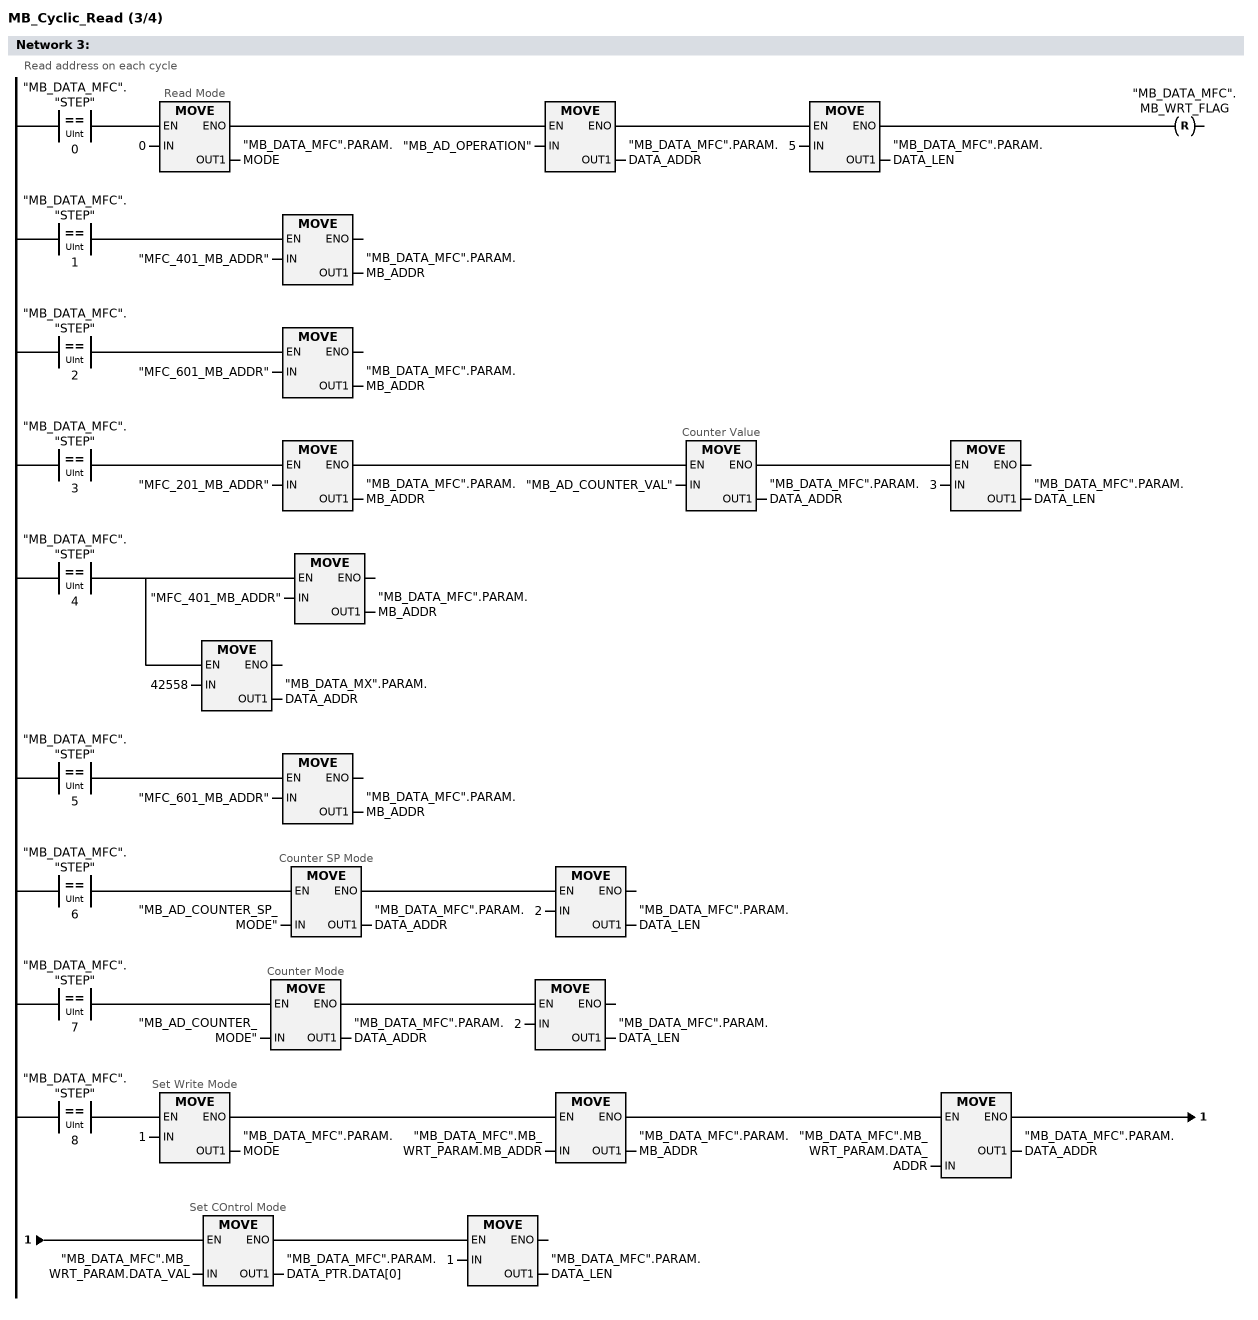
   RUNG wire#powerrail
      { S7_Templates := "SrcType := UInt" } EQ_Contact(in1 := "MB_DATA_MFC"."STEP", in2 := 0)
      Move(in := 0, out1 => "MB_DATA_MFC".PARAM.MODE)   // Read Mode
      Move(in := "MB_AD_OPERATION", out1 => "MB_DATA_MFC".PARAM.DATA_ADDR)
      Move(in := 5, out1 => "MB_DATA_MFC".PARAM.DATA_LEN)
      R_Coil( "MB_DATA_MFC".MB_WRT_FLAG )
   END_RUNG
   RUNG wire#powerrail
      { S7_Templates := "SrcType := UInt" } EQ_Contact(in1 := "MB_DATA_MFC"."STEP", in2 := 1)
      Move(in := "MFC_401_MB_ADDR", out1 => "MB_DATA_MFC".PARAM.MB_ADDR)
   END_RUNG
   RUNG wire#powerrail
      { S7_Templates := "SrcType := UInt" } EQ_Contact(in1 := "MB_DATA_MFC"."STEP", in2 := 2)
      Move(in := "MFC_601_MB_ADDR", out1 => "MB_DATA_MFC".PARAM.MB_ADDR)
   END_RUNG
   RUNG wire#powerrail
      { S7_Templates := "SrcType := UInt" } EQ_Contact(in1 := "MB_DATA_MFC"."STEP", in2 := 3)
      Move(in := "MFC_201_MB_ADDR", out1 => "MB_DATA_MFC".PARAM.MB_ADDR)
      Move(in := "MB_AD_COUNTER_VAL", out1 => "MB_DATA_MFC".PARAM.DATA_ADDR)   // Counter Value
      Move(in := 3, out1 => "MB_DATA_MFC".PARAM.DATA_LEN)
   END_RUNG
   RUNG wire#powerrail
      { S7_Templates := "SrcType := UInt" } EQ_Contact(in1 := "MB_DATA_MFC"."STEP", in2 := 4)
      wire#w1
      Move(in := "MFC_401_MB_ADDR", out1 => "MB_DATA_MFC".PARAM.MB_ADDR)
   END_RUNG
   RUNG wire#w1
      Move(in := 42558, out1 => "MB_DATA_MX".PARAM.DATA_ADDR)
   END_RUNG
   RUNG wire#powerrail
      { S7_Templates := "SrcType := UInt" } EQ_Contact(in1 := "MB_DATA_MFC"."STEP", in2 := 5)
      Move(in := "MFC_601_MB_ADDR", out1 => "MB_DATA_MFC".PARAM.MB_ADDR)
   END_RUNG
   RUNG wire#powerrail
      { S7_Templates := "SrcType := UInt" } EQ_Contact(in1 := "MB_DATA_MFC"."STEP", in2 := 6)
      Move(in := "MB_AD_COUNTER_SP_MODE", out1 => "MB_DATA_MFC".PARAM.DATA_ADDR)   // Counter SP Mode
      Move(in := 2, out1 => "MB_DATA_MFC".PARAM.DATA_LEN)
   END_RUNG
   RUNG wire#powerrail
      { S7_Templates := "SrcType := UInt" } EQ_Contact(in1 := "MB_DATA_MFC"."STEP", in2 := 7)
      Move(in := "MB_AD_COUNTER_MODE", out1 => "MB_DATA_MFC".PARAM.DATA_ADDR)   // Counter Mode
      Move(in := 2, out1 => "MB_DATA_MFC".PARAM.DATA_LEN)
   END_RUNG
   RUNG wire#powerrail
      { S7_Templates := "SrcType := UInt" } EQ_Contact(in1 := "MB_DATA_MFC"."STEP", in2 := 8)
      Move(in := 1, out1 => "MB_DATA_MFC".PARAM.MODE)   // Set Write Mode
      Move(in := "MB_DATA_MFC".MB_WRT_PARAM.MB_ADDR, out1 => "MB_DATA_MFC".PARAM.MB_ADDR)
      Move(in := "MB_DATA_MFC".MB_WRT_PARAM.DATA_ADDR, out1 => "MB_DATA_MFC".PARAM.DATA_ADDR)
      Move(in := "MB_DATA_MFC".MB_WRT_PARAM.DATA_VAL, out1 => "MB_DATA_MFC".PARAM.DATA_PTR.DATA[0])   // Set COntrol Mode
      Move(in := 1, out1 => "MB_DATA_MFC".PARAM.DATA_LEN)
   END_RUNG
   // the same network as SCL:
   IF "MB_DATA_MFC"."STEP" = 0 THEN
       "MB_DATA_MFC".PARAM.MODE := 0;   // Read Mode
       "MB_DATA_MFC".PARAM.DATA_ADDR := "MB_AD_OPERATION";
       "MB_DATA_MFC".PARAM.DATA_LEN := 5;
       "MB_DATA_MFC".MB_WRT_FLAG := FALSE;
   END_IF;
   IF "MB_DATA_MFC"."STEP" = 1 THEN "MB_DATA_MFC".PARAM.MB_ADDR := "MFC_401_MB_ADDR"; END_IF;
   IF "MB_DATA_MFC"."STEP" = 2 THEN "MB_DATA_MFC".PARAM.MB_ADDR := "MFC_601_MB_ADDR"; END_IF;
   IF "MB_DATA_MFC"."STEP" = 3 THEN
       "MB_DATA_MFC".PARAM.MB_ADDR := "MFC_201_MB_ADDR";
       "MB_DATA_MFC".PARAM.DATA_ADDR := "MB_AD_COUNTER_VAL";   // Counter Value
       "MB_DATA_MFC".PARAM.DATA_LEN := 3;
   END_IF;
   IF "MB_DATA_MFC"."STEP" = 4 THEN
       "MB_DATA_MFC".PARAM.MB_ADDR := "MFC_401_MB_ADDR";
       "MB_DATA_MX".PARAM.DATA_ADDR := 42558;
   END_IF;
   IF "MB_DATA_MFC"."STEP" = 5 THEN "MB_DATA_MFC".PARAM.MB_ADDR := "MFC_601_MB_ADDR"; END_IF;
   IF "MB_DATA_MFC"."STEP" = 6 THEN
       "MB_DATA_MFC".PARAM.DATA_ADDR := "MB_AD_COUNTER_SP_MODE";   // Counter SP Mode
       "MB_DATA_MFC".PARAM.DATA_LEN := 2;
   END_IF;
   IF "MB_DATA_MFC"."STEP" = 7 THEN
       "MB_DATA_MFC".PARAM.DATA_ADDR := "MB_AD_COUNTER_MODE";   // Counter Mode
       "MB_DATA_MFC".PARAM.DATA_LEN := 2;
   END_IF;
   IF "MB_DATA_MFC"."STEP" = 8 THEN
       "MB_DATA_MFC".PARAM.MODE := 1;   // Set Write Mode
       "MB_DATA_MFC".PARAM.MB_ADDR := "MB_DATA_MFC".MB_WRT_PARAM.MB_ADDR;
       "MB_DATA_MFC".PARAM.DATA_ADDR := "MB_DATA_MFC".MB_WRT_PARAM.DATA_ADDR;
       "MB_DATA_MFC".PARAM.DATA_PTR.DATA[0] := "MB_DATA_MFC".MB_WRT_PARAM.DATA_VAL;   // Set COntrol Mode
       "MB_DATA_MFC".PARAM.DATA_LEN := 1;
   END_IF;
END_REGION

REGION Network 4
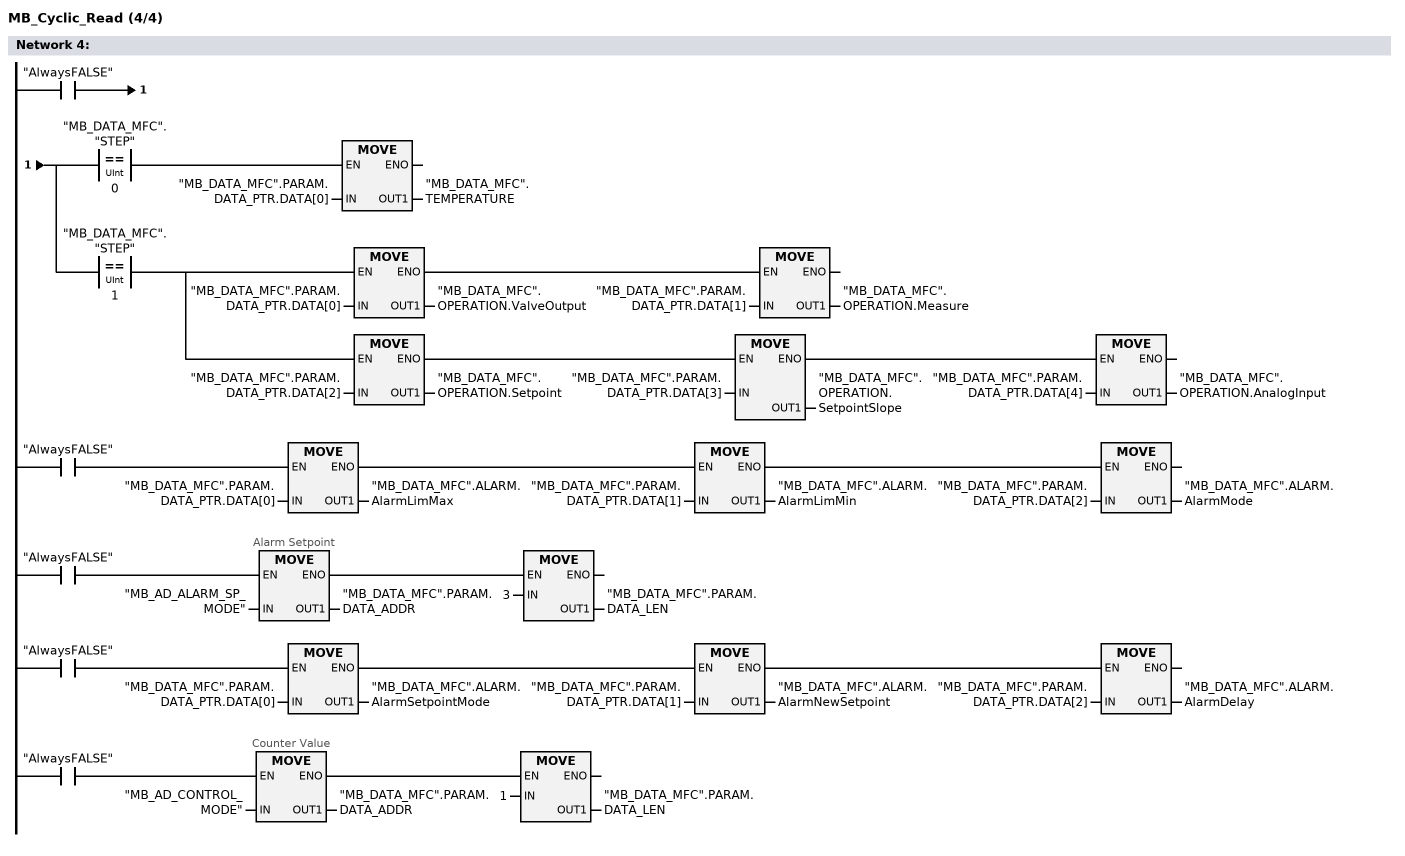
   RUNG wire#powerrail
      Contact( "AlwaysFALSE" )
      wire#w1
      { S7_Templates := "SrcType := UInt" } EQ_Contact(in1 := "MB_DATA_MFC"."STEP", in2 := 0)
      Move(in := "MB_DATA_MFC".PARAM.DATA_PTR.DATA[0], out1 => "MB_DATA_MFC".TEMPERATURE)
   END_RUNG
   RUNG wire#w1
      { S7_Templates := "SrcType := UInt" } EQ_Contact(in1 := "MB_DATA_MFC"."STEP", in2 := 1)
      wire#w2
      Move(in := "MB_DATA_MFC".PARAM.DATA_PTR.DATA[0], out1 => "MB_DATA_MFC".OPERATION.ValveOutput)
      Move(in := "MB_DATA_MFC".PARAM.DATA_PTR.DATA[1], out1 => "MB_DATA_MFC".OPERATION.Measure)
   END_RUNG
   RUNG wire#w2
      Move(in := "MB_DATA_MFC".PARAM.DATA_PTR.DATA[2], out1 => "MB_DATA_MFC".OPERATION.Setpoint)
      Move(in := "MB_DATA_MFC".PARAM.DATA_PTR.DATA[3], out1 => "MB_DATA_MFC".OPERATION.SetpointSlope)
      Move(in := "MB_DATA_MFC".PARAM.DATA_PTR.DATA[4], out1 => "MB_DATA_MFC".OPERATION.AnalogInput)
   END_RUNG
   RUNG wire#powerrail
      Contact( "AlwaysFALSE" )
      Move(in := "MB_DATA_MFC".PARAM.DATA_PTR.DATA[0], out1 => "MB_DATA_MFC".ALARM.AlarmLimMax)
      Move(in := "MB_DATA_MFC".PARAM.DATA_PTR.DATA[1], out1 => "MB_DATA_MFC".ALARM.AlarmLimMin)
      Move(in := "MB_DATA_MFC".PARAM.DATA_PTR.DATA[2], out1 => "MB_DATA_MFC".ALARM.AlarmMode)
   END_RUNG
   RUNG wire#powerrail
      Contact( "AlwaysFALSE" )
      Move(in := "MB_AD_ALARM_SP_MODE", out1 => "MB_DATA_MFC".PARAM.DATA_ADDR)   // Alarm Setpoint
      Move(in := 3, out1 => "MB_DATA_MFC".PARAM.DATA_LEN)
   END_RUNG
   RUNG wire#powerrail
      Contact( "AlwaysFALSE" )
      Move(in := "MB_DATA_MFC".PARAM.DATA_PTR.DATA[0], out1 => "MB_DATA_MFC".ALARM.AlarmSetpointMode)
      Move(in := "MB_DATA_MFC".PARAM.DATA_PTR.DATA[1], out1 => "MB_DATA_MFC".ALARM.AlarmNewSetpoint)
      Move(in := "MB_DATA_MFC".PARAM.DATA_PTR.DATA[2], out1 => "MB_DATA_MFC".ALARM.AlarmDelay)
   END_RUNG
   RUNG wire#powerrail
      Contact( "AlwaysFALSE" )
      Move(in := "MB_AD_CONTROL_MODE", out1 => "MB_DATA_MFC".PARAM.DATA_ADDR)   // Counter Value
      Move(in := 1, out1 => "MB_DATA_MFC".PARAM.DATA_LEN)
   END_RUNG
   // the same network as SCL:
   IF "AlwaysFALSE" AND ("MB_DATA_MFC"."STEP" = 0) THEN
       "MB_DATA_MFC".TEMPERATURE := "MB_DATA_MFC".PARAM.DATA_PTR.DATA[0];
   END_IF;
   IF "AlwaysFALSE" AND ("MB_DATA_MFC"."STEP" = 1) THEN
       "MB_DATA_MFC".OPERATION.ValveOutput := "MB_DATA_MFC".PARAM.DATA_PTR.DATA[0];
       "MB_DATA_MFC".OPERATION.Measure := "MB_DATA_MFC".PARAM.DATA_PTR.DATA[1];
       "MB_DATA_MFC".OPERATION.Setpoint := "MB_DATA_MFC".PARAM.DATA_PTR.DATA[2];
       "MB_DATA_MFC".OPERATION.SetpointSlope := "MB_DATA_MFC".PARAM.DATA_PTR.DATA[3];
       "MB_DATA_MFC".OPERATION.AnalogInput := "MB_DATA_MFC".PARAM.DATA_PTR.DATA[4];
   END_IF;
   IF "AlwaysFALSE" THEN
       "MB_DATA_MFC".ALARM.AlarmLimMax := "MB_DATA_MFC".PARAM.DATA_PTR.DATA[0];
       "MB_DATA_MFC".ALARM.AlarmLimMin := "MB_DATA_MFC".PARAM.DATA_PTR.DATA[1];
       "MB_DATA_MFC".ALARM.AlarmMode := "MB_DATA_MFC".PARAM.DATA_PTR.DATA[2];
       "MB_DATA_MFC".PARAM.DATA_ADDR := "MB_AD_ALARM_SP_MODE";   // Alarm Setpoint
       "MB_DATA_MFC".PARAM.DATA_LEN := 3;
       "MB_DATA_MFC".ALARM.AlarmSetpointMode := "MB_DATA_MFC".PARAM.DATA_PTR.DATA[0];
       "MB_DATA_MFC".ALARM.AlarmNewSetpoint := "MB_DATA_MFC".PARAM.DATA_PTR.DATA[1];
       "MB_DATA_MFC".ALARM.AlarmDelay := "MB_DATA_MFC".PARAM.DATA_PTR.DATA[2];
       "MB_DATA_MFC".PARAM.DATA_ADDR := "MB_AD_CONTROL_MODE";   // Counter Value
       "MB_DATA_MFC".PARAM.DATA_LEN := 1;
   END_IF;
END_REGION
END_FUNCTION

FUNCTION "TESTS_1" : Void   // FC13, LAD
{ S7_Optimized_Access := 'FALSE' }
VERSION : 0.1
   VAR_TEMP   // added for the SCL form of the ladder/FBD networks
      _w1 : Bool;
   END_VAR
BEGIN

REGION Network 1
   // ALARM Settings
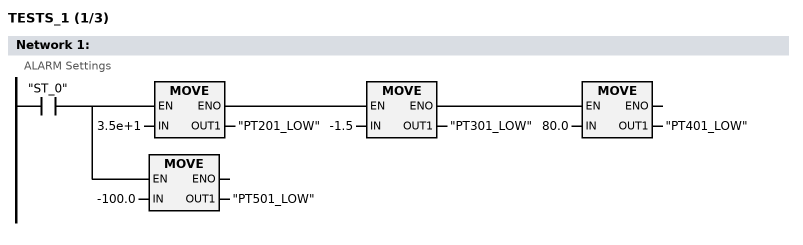
   RUNG wire#powerrail
      Contact( "ST_0" )
      wire#w1
      { S7_GenerateENO := "TRUE" } Move(in := 3.5e+1, out1 => "PT201_LOW")
      { S7_GenerateENO := "TRUE" } Move(in := -1.5, out1 => "PT301_LOW")
      { S7_GenerateENO := "TRUE" } Move(in := 80.0, out1 => "PT401_LOW")
   END_RUNG
   RUNG wire#w1
      { S7_GenerateENO := "TRUE" } Move(in := -100.0, out1 => "PT501_LOW")
   END_RUNG
   // the same network as SCL:
   // ENO of a box is taken as its EN; it also drops when the box reports an error
   IF "ST_0" THEN
       "PT201_LOW" := 3.5e+1;
       "PT301_LOW" := -1.5;
       "PT401_LOW" := 80.0;
       "PT501_LOW" := -100.0;
   END_IF;
END_REGION

REGION Network 2: Pneumatic Tests
   // Test Pneumatic System (Test #1-#6)
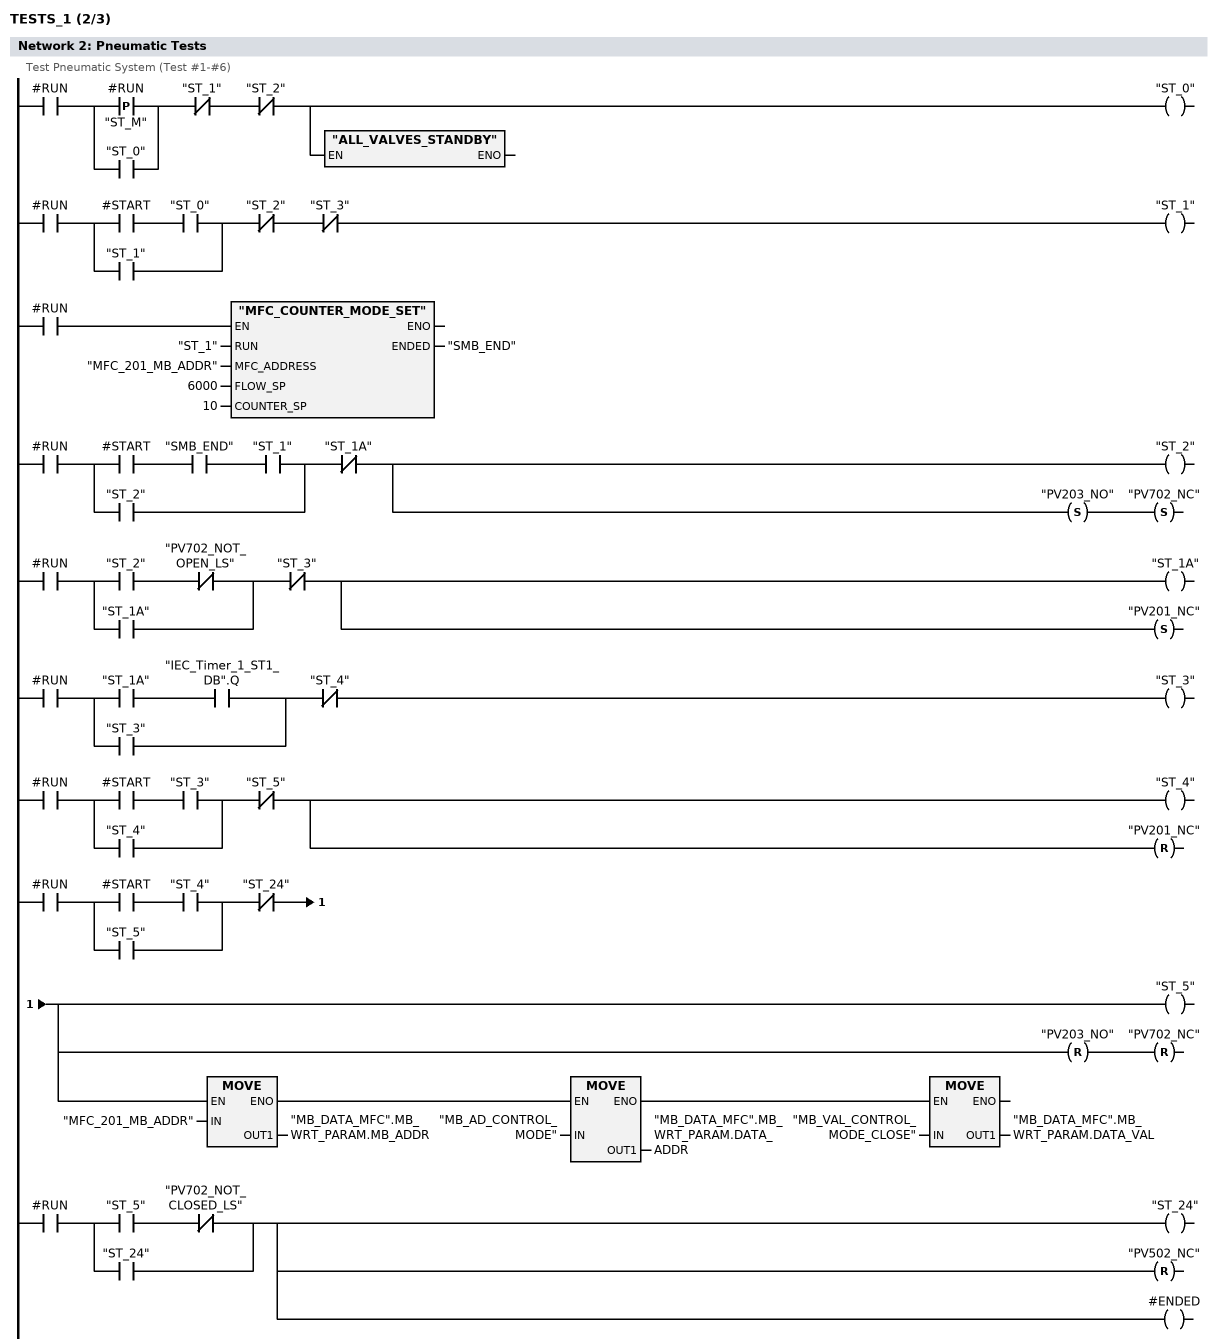
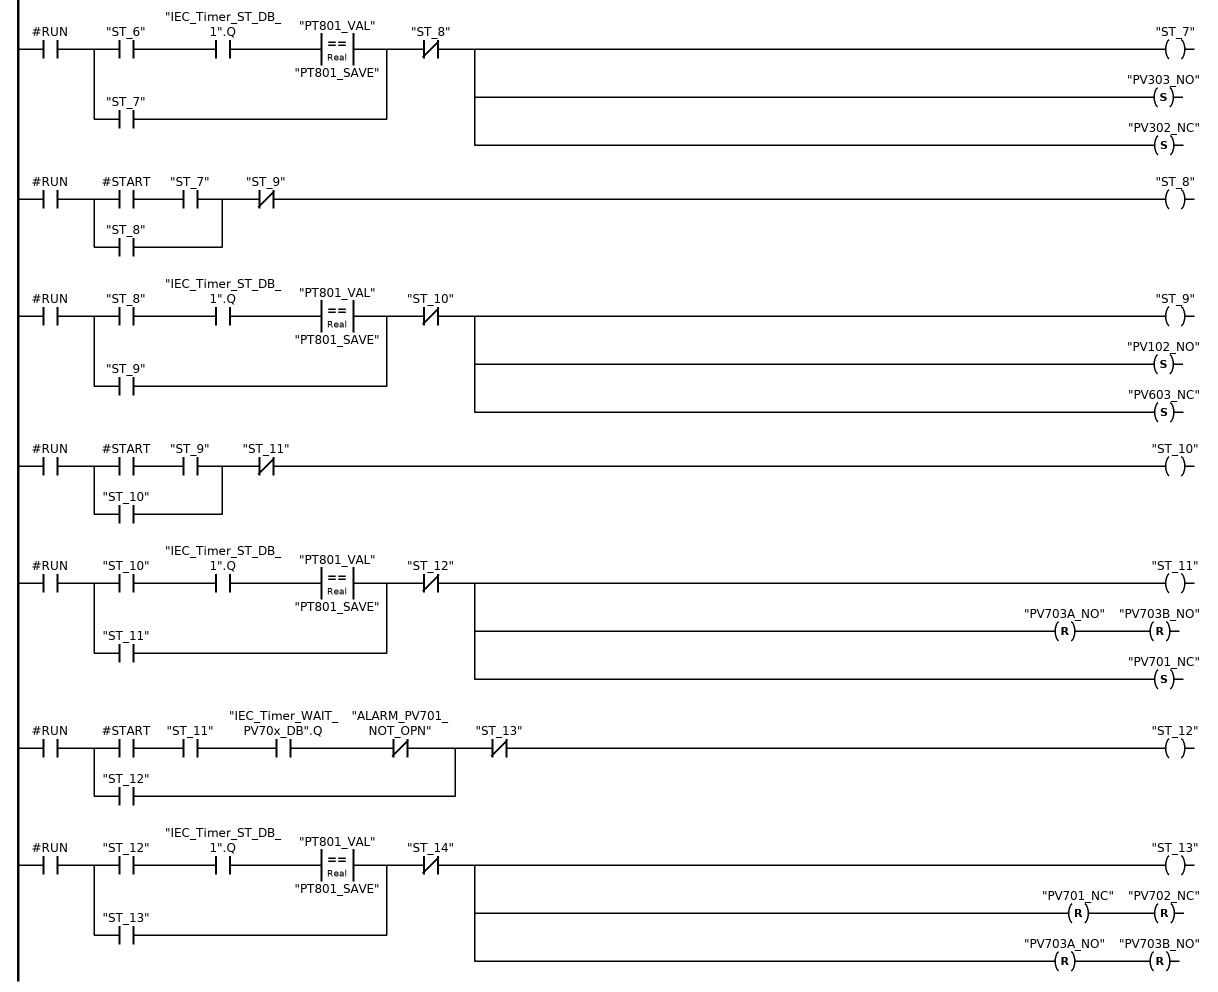
   RUNG wire#powerrail
      Contact( #RUN )
      wire#w1
      P_Contact(operand := #RUN, bit := "ST_M")
      wire#w2
      I_Contact( "ST_1" )
      I_Contact( "ST_2" )
      wire#w3
      Coil( "ST_0" )
   END_RUNG
   RUNG wire#w1
      Contact( "ST_0" )
   END_RUNG wire#w2
   RUNG wire#w3
      "ALL_VALVES_STANDBY"()
   END_RUNG
   RUNG wire#powerrail
      Contact( #RUN )
      wire#w4
      Contact( #START )
      Contact( "ST_0" )
      wire#w5
      I_Contact( "ST_2" )
      I_Contact( "ST_3" )
      Coil( "ST_1" )
   END_RUNG
   RUNG wire#w4
      Contact( "ST_1" )
   END_RUNG wire#w5
   RUNG wire#powerrail
      Contact( #RUN )
      "MFC_COUNTER_MODE_SET"(RUN := "ST_1", MFC_ADDRESS := "MFC_201_MB_ADDR", FLOW_SP := 6000, COUNTER_SP := 10, ENDED => "SMB_END")
   END_RUNG
   RUNG wire#powerrail
      Contact( #RUN )
      wire#w6
      Contact( #START )
      Contact( "SMB_END" )
      Contact( "ST_1" )
      wire#w7
      I_Contact( "ST_1A" )
      wire#w8
      Coil( "ST_2" )
   END_RUNG
   RUNG wire#w6
      Contact( "ST_2" )
   END_RUNG wire#w7
   RUNG wire#w8
      S_Coil( "PV203_NO" )
      S_Coil( "PV702_NC" )
   END_RUNG
   RUNG wire#powerrail
      Contact( #RUN )
      wire#w9
      Contact( "ST_2" )
      I_Contact( "PV702_NOT_OPEN_LS" )
      wire#w10
      I_Contact( "ST_3" )
      wire#w11
      Coil( "ST_1A" )
   END_RUNG
   RUNG wire#w9
      Contact( "ST_1A" )
   END_RUNG wire#w10
   RUNG wire#w11
      S_Coil( "PV201_NC" )
   END_RUNG
   RUNG wire#powerrail
      Contact( #RUN )
      wire#w12
      Contact( "ST_1A" )
      Contact( "IEC_Timer_1_ST1_DB".Q )
      wire#w13
      I_Contact( "ST_4" )
      Coil( "ST_3" )
   END_RUNG
   RUNG wire#w12
      Contact( "ST_3" )
   END_RUNG wire#w13
   RUNG wire#powerrail
      Contact( #RUN )
      wire#w14
      Contact( #START )
      Contact( "ST_3" )
      wire#w15
      I_Contact( "ST_5" )
      wire#w16
      Coil( "ST_4" )
   END_RUNG
   RUNG wire#w14
      Contact( "ST_4" )
   END_RUNG wire#w15
   RUNG wire#w16
      R_Coil( "PV201_NC" )
   END_RUNG
   RUNG wire#powerrail
      Contact( #RUN )
      wire#w17
      Contact( #START )
      Contact( "ST_4" )
      wire#w18
      I_Contact( "ST_24" )
      wire#w19
      Coil( "ST_5" )
   END_RUNG
   RUNG wire#w17
      Contact( "ST_5" )
   END_RUNG wire#w18
   RUNG wire#w19
      R_Coil( "PV203_NO" )
      R_Coil( "PV702_NC" )
   END_RUNG
   RUNG wire#w19
      Move(in := "MFC_201_MB_ADDR", out1 => "MB_DATA_MFC".MB_WRT_PARAM.MB_ADDR)
      Move(in := "MB_AD_CONTROL_MODE", out1 => "MB_DATA_MFC".MB_WRT_PARAM.DATA_ADDR)
      Move(in := "MB_VAL_CONTROL_MODE_CLOSE", out1 => "MB_DATA_MFC".MB_WRT_PARAM.DATA_VAL)
   END_RUNG
   RUNG wire#powerrail
      Contact( #RUN )
      wire#w20
      Contact( "ST_5" )
      I_Contact( "PV702_NOT_CLOSED_LS" )
      wire#w21
      Coil( "ST_24" )
   END_RUNG
   RUNG wire#w20
      Contact( "ST_24" )
   END_RUNG wire#w21
   RUNG wire#w21
      R_Coil( "PV502_NC" )
   END_RUNG
   RUNG wire#w21
      Coil( #ENDED )
   END_RUNG
   RUNG wire#powerrail
      Contact( #RUN )
      wire#w22
      Contact( "ST_6" )
      Contact( "IEC_Timer_ST_DB_1".Q )
      { S7_Templates := "SrcType := Real" } EQ_Contact(in1 := "PT801_VAL", in2 := "PT801_SAVE")
      wire#w23
      I_Contact( "ST_8" )
      wire#w24
      Coil( "ST_7" )
   END_RUNG
   RUNG wire#w22
      Contact( "ST_7" )
   END_RUNG wire#w23
   RUNG wire#w24
      S_Coil( "PV303_NO" )
   END_RUNG
   RUNG wire#w24
      S_Coil( "PV302_NC" )
   END_RUNG
   RUNG wire#powerrail
      Contact( #RUN )
      wire#w25
      Contact( #START )
      Contact( "ST_7" )
      wire#w26
      I_Contact( "ST_9" )
      Coil( "ST_8" )
   END_RUNG
   RUNG wire#w25
      Contact( "ST_8" )
   END_RUNG wire#w26
   RUNG wire#powerrail
      Contact( #RUN )
      wire#w27
      Contact( "ST_8" )
      Contact( "IEC_Timer_ST_DB_1".Q )
      { S7_Templates := "SrcType := Real" } EQ_Contact(in1 := "PT801_VAL", in2 := "PT801_SAVE")
      wire#w28
      I_Contact( "ST_10" )
      wire#w29
      Coil( "ST_9" )
   END_RUNG
   RUNG wire#w27
      Contact( "ST_9" )
   END_RUNG wire#w28
   RUNG wire#w29
      S_Coil( "PV102_NO" )
   END_RUNG
   RUNG wire#w29
      S_Coil( "PV603_NC" )
   END_RUNG
   RUNG wire#powerrail
      Contact( #RUN )
      wire#w30
      Contact( #START )
      Contact( "ST_9" )
      wire#w31
      I_Contact( "ST_11" )
      Coil( "ST_10" )
   END_RUNG
   RUNG wire#w30
      Contact( "ST_10" )
   END_RUNG wire#w31
   RUNG wire#powerrail
      Contact( #RUN )
      wire#w32
      Contact( "ST_10" )
      Contact( "IEC_Timer_ST_DB_1".Q )
      { S7_Templates := "SrcType := Real" } EQ_Contact(in1 := "PT801_VAL", in2 := "PT801_SAVE")
      wire#w33
      I_Contact( "ST_12" )
      wire#w34
      Coil( "ST_11" )
   END_RUNG
   RUNG wire#w32
      Contact( "ST_11" )
   END_RUNG wire#w33
   RUNG wire#w34
      R_Coil( "PV703A_NO" )
      R_Coil( "PV703B_NO" )
   END_RUNG
   RUNG wire#w34
      S_Coil( "PV701_NC" )
   END_RUNG
   RUNG wire#powerrail
      Contact( #RUN )
      wire#w35
      Contact( #START )
      Contact( "ST_11" )
      Contact( "IEC_Timer_WAIT_PV70x_DB".Q )
      I_Contact( "ALARM_PV701_NOT_OPN" )
      wire#w36
      I_Contact( "ST_13" )
      Coil( "ST_12" )
   END_RUNG
   RUNG wire#w35
      Contact( "ST_12" )
   END_RUNG wire#w36
   RUNG wire#powerrail
      Contact( #RUN )
      wire#w37
      Contact( "ST_12" )
      Contact( "IEC_Timer_ST_DB_1".Q )
      { S7_Templates := "SrcType := Real" } EQ_Contact(in1 := "PT801_VAL", in2 := "PT801_SAVE")
      wire#w38
      I_Contact( "ST_14" )
      wire#w39
      Coil( "ST_13" )
   END_RUNG
   RUNG wire#w37
      Contact( "ST_13" )
   END_RUNG wire#w38
   RUNG wire#w39
      R_Coil( "PV701_NC" )
      R_Coil( "PV702_NC" )
   END_RUNG
   RUNG wire#w39
      R_Coil( "PV703A_NO" )
      R_Coil( "PV703B_NO" )
   END_RUNG
   // the same network as SCL:
   #_w1 := #RUN AND #RUN AND NOT "ST_M";   // rising edge of #RUN
   "ST_M" := #RUN;
   "ST_0" := (#_w1 OR (#RUN AND "ST_0")) AND NOT "ST_1" AND NOT "ST_2";
   IF "ST_0" THEN "ALL_VALVES_STANDBY"(); END_IF;
   "ST_1" := #RUN AND ((#START AND "ST_0") OR "ST_1") AND NOT "ST_2" AND NOT "ST_3";
   IF #RUN THEN
       "MFC_COUNTER_MODE_SET"(RUN := "ST_1",
                              MFC_ADDRESS := "MFC_201_MB_ADDR",
                              FLOW_SP := 6000,
                              COUNTER_SP := 10,
                              ENDED => "SMB_END");
   END_IF;
   "ST_2" := #RUN AND ((#START AND "SMB_END" AND "ST_1") OR "ST_2") AND NOT "ST_1A";
   IF "ST_2" THEN
       "PV203_NO" := TRUE;
       "PV702_NC" := TRUE;
   END_IF;
   "ST_1A" := #RUN AND (("ST_2" AND NOT "PV702_NOT_OPEN_LS") OR "ST_1A") AND NOT "ST_3";
   IF "ST_1A" THEN "PV201_NC" := TRUE; END_IF;
   "ST_3" := #RUN AND (("ST_1A" AND "IEC_Timer_1_ST1_DB".Q) OR "ST_3") AND NOT "ST_4";
   "ST_4" := #RUN AND ((#START AND "ST_3") OR "ST_4") AND NOT "ST_5";
   IF "ST_4" THEN "PV201_NC" := FALSE; END_IF;
   "ST_5" := #RUN AND ((#START AND "ST_4") OR "ST_5") AND NOT "ST_24";
   IF "ST_5" THEN
       "PV203_NO" := FALSE;
       "PV702_NC" := FALSE;
       "MB_DATA_MFC".MB_WRT_PARAM.MB_ADDR := "MFC_201_MB_ADDR";
       "MB_DATA_MFC".MB_WRT_PARAM.DATA_ADDR := "MB_AD_CONTROL_MODE";
       "MB_DATA_MFC".MB_WRT_PARAM.DATA_VAL := "MB_VAL_CONTROL_MODE_CLOSE";
   END_IF;
   "ST_24" := #RUN AND (("ST_5" AND NOT "PV702_NOT_CLOSED_LS") OR "ST_24");
   IF "ST_24" THEN "PV502_NC" := FALSE; END_IF;
   #ENDED := "ST_24";
   "ST_7" := #RUN AND (("ST_6" AND "IEC_Timer_ST_DB_1".Q AND ("PT801_VAL" = "PT801_SAVE")) OR "ST_7") AND NOT "ST_8";
   IF "ST_7" THEN
       "PV303_NO" := TRUE;
       "PV302_NC" := TRUE;
   END_IF;
   "ST_8" := #RUN AND ((#START AND "ST_7") OR "ST_8") AND NOT "ST_9";
   "ST_9" := #RUN AND (("ST_8" AND "IEC_Timer_ST_DB_1".Q AND ("PT801_VAL" = "PT801_SAVE")) OR "ST_9") AND NOT "ST_10";
   IF "ST_9" THEN
       "PV102_NO" := TRUE;
       "PV603_NC" := TRUE;
   END_IF;
   "ST_10" := #RUN AND ((#START AND "ST_9") OR "ST_10") AND NOT "ST_11";
   "ST_11" := #RUN AND (("ST_10" AND "IEC_Timer_ST_DB_1".Q AND ("PT801_VAL" = "PT801_SAVE")) OR "ST_11") AND NOT "ST_12";
   IF "ST_11" THEN
       "PV703A_NO" := FALSE;
       "PV703B_NO" := FALSE;
       "PV701_NC" := TRUE;
   END_IF;
   "ST_12" := #RUN AND ((#START AND "ST_11" AND "IEC_Timer_WAIT_PV70x_DB".Q AND NOT "ALARM_PV701_NOT_OPN") OR "ST_12") AND NOT "ST_13";
   "ST_13" := #RUN AND (("ST_12" AND "IEC_Timer_ST_DB_1".Q AND ("PT801_VAL" = "PT801_SAVE")) OR "ST_13") AND NOT "ST_14";
   IF "ST_13" THEN
       "PV701_NC" := FALSE;
       "PV702_NC" := FALSE;
       "PV703A_NO" := FALSE;
       "PV703B_NO" := FALSE;
   END_IF;
END_REGION

REGION Network 3: Process Tests
   // Tests Process Circuits  (Test #7-#9)
END_REGION

REGION Network 4
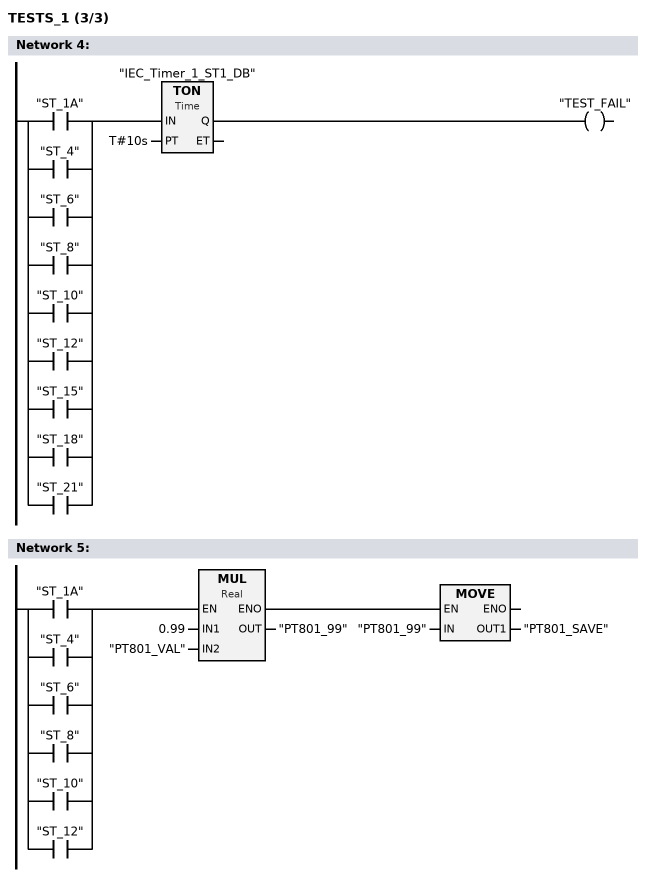
   "IEC_Timer_1_ST1_DB".TON(IN := "ST_1A" OR "ST_4" OR "ST_6" OR "ST_8" OR "ST_10" OR "ST_12" OR "ST_15" OR "ST_18" OR "ST_21",
                           PT := T#10s);
   "TEST_FAIL" := "IEC_Timer_1_ST1_DB".Q;
END_REGION

REGION Network 5
   RUNG wire#powerrail
      Contact( "ST_1A" )
      wire#w1
      { S7_Templates := "SrcType := Real" } Mul(in1 := 0.99, in2 := "PT801_VAL", out => "PT801_99")
      { S7_GenerateENO := "TRUE" } Move(in := "PT801_99", out1 => "PT801_SAVE")
   END_RUNG
   RUNG wire#powerrail
      Contact( "ST_4" )
   END_RUNG wire#w1
   RUNG wire#powerrail
      Contact( "ST_6" )
   END_RUNG wire#w1
   RUNG wire#powerrail
      Contact( "ST_8" )
   END_RUNG wire#w1
   RUNG wire#powerrail
      Contact( "ST_10" )
   END_RUNG wire#w1
   RUNG wire#powerrail
      Contact( "ST_12" )
   END_RUNG wire#w1
   // the same network as SCL:
   IF "ST_1A" OR "ST_4" OR "ST_6" OR "ST_8" OR "ST_10" OR "ST_12" THEN
       "PT801_99" := 0.99 * "PT801_VAL";
       "PT801_SAVE" := "PT801_99";
   END_IF;
END_REGION
END_FUNCTION

FUNCTION "ALARMS" : Void   // FC14, LAD
{ S7_Optimized_Access := 'FALSE' }
VERSION : 0.1
// Removed Doors Alarm
BEGIN

REGION Network 1
   // LOW ALARMS
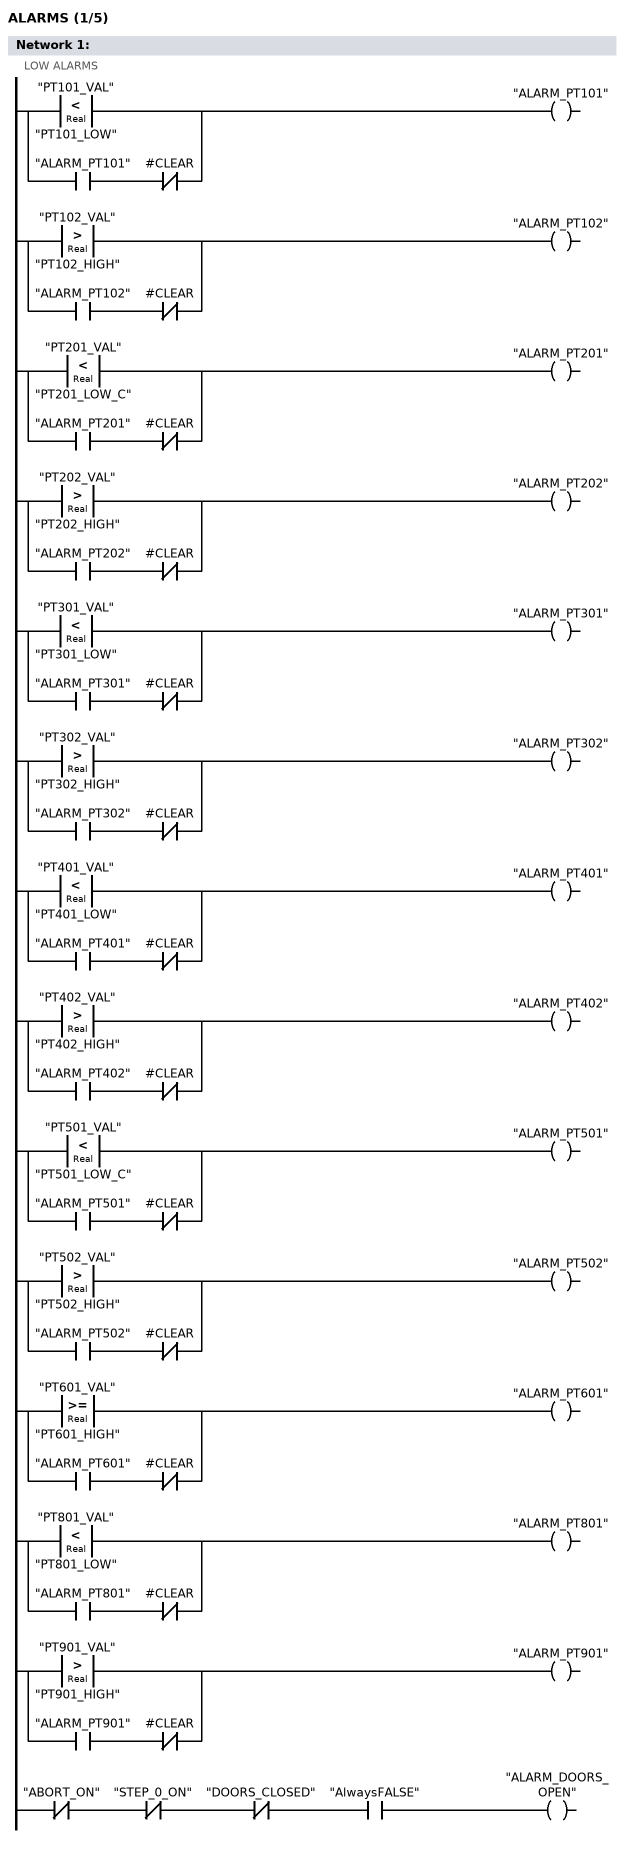
   RUNG wire#powerrail
      { S7_Templates := "SrcType := Real" } LT_Contact(in1 := "PT101_VAL", in2 := "PT101_LOW")
      wire#w1
      Coil( "ALARM_PT101" )
   END_RUNG
   RUNG wire#powerrail
      Contact( "ALARM_PT101" )
      I_Contact( #CLEAR )
   END_RUNG wire#w1
   RUNG wire#powerrail
      { S7_Templates := "SrcType := Real" } GT_Contact(in1 := "PT102_VAL", in2 := "PT102_HIGH")
      wire#w2
      Coil( "ALARM_PT102" )
   END_RUNG
   RUNG wire#powerrail
      Contact( "ALARM_PT102" )
      I_Contact( #CLEAR )
   END_RUNG wire#w2
   RUNG wire#powerrail
      { S7_Templates := "SrcType := Real" } LT_Contact(in1 := "PT201_VAL", in2 := "PT201_LOW_C")
      wire#w3
      Coil( "ALARM_PT201" )
   END_RUNG
   RUNG wire#powerrail
      Contact( "ALARM_PT201" )
      I_Contact( #CLEAR )
   END_RUNG wire#w3
   RUNG wire#powerrail
      { S7_Templates := "SrcType := Real" } GT_Contact(in1 := "PT202_VAL", in2 := "PT202_HIGH")
      wire#w4
      Coil( "ALARM_PT202" )
   END_RUNG
   RUNG wire#powerrail
      Contact( "ALARM_PT202" )
      I_Contact( #CLEAR )
   END_RUNG wire#w4
   RUNG wire#powerrail
      { S7_Templates := "SrcType := Real" } LT_Contact(in1 := "PT301_VAL", in2 := "PT301_LOW")
      wire#w5
      Coil( "ALARM_PT301" )
   END_RUNG
   RUNG wire#powerrail
      Contact( "ALARM_PT301" )
      I_Contact( #CLEAR )
   END_RUNG wire#w5
   RUNG wire#powerrail
      { S7_Templates := "SrcType := Real" } GT_Contact(in1 := "PT302_VAL", in2 := "PT302_HIGH")
      wire#w6
      Coil( "ALARM_PT302" )
   END_RUNG
   RUNG wire#powerrail
      Contact( "ALARM_PT302" )
      I_Contact( #CLEAR )
   END_RUNG wire#w6
   RUNG wire#powerrail
      { S7_Templates := "SrcType := Real" } LT_Contact(in1 := "PT401_VAL", in2 := "PT401_LOW")
      wire#w7
      Coil( "ALARM_PT401" )
   END_RUNG
   RUNG wire#powerrail
      Contact( "ALARM_PT401" )
      I_Contact( #CLEAR )
   END_RUNG wire#w7
   RUNG wire#powerrail
      { S7_Templates := "SrcType := Real" } GT_Contact(in1 := "PT402_VAL", in2 := "PT402_HIGH")
      wire#w8
      Coil( "ALARM_PT402" )
   END_RUNG
   RUNG wire#powerrail
      Contact( "ALARM_PT402" )
      I_Contact( #CLEAR )
   END_RUNG wire#w8
   RUNG wire#powerrail
      { S7_Templates := "SrcType := Real" } LT_Contact(in1 := "PT501_VAL", in2 := "PT501_LOW_C")
      wire#w9
      Coil( "ALARM_PT501" )
   END_RUNG
   RUNG wire#powerrail
      Contact( "ALARM_PT501" )
      I_Contact( #CLEAR )
   END_RUNG wire#w9
   RUNG wire#powerrail
      { S7_Templates := "SrcType := Real" } GT_Contact(in1 := "PT502_VAL", in2 := "PT502_HIGH")
      wire#w10
      Coil( "ALARM_PT502" )
   END_RUNG
   RUNG wire#powerrail
      Contact( "ALARM_PT502" )
      I_Contact( #CLEAR )
   END_RUNG wire#w10
   RUNG wire#powerrail
      { S7_Templates := "SrcType := Real" } GE_Contact(in1 := "PT601_VAL", in2 := "PT601_HIGH")
      wire#w11
      Coil( "ALARM_PT601" )
   END_RUNG
   RUNG wire#powerrail
      Contact( "ALARM_PT601" )
      I_Contact( #CLEAR )
   END_RUNG wire#w11
   RUNG wire#powerrail
      { S7_Templates := "SrcType := Real" } LT_Contact(in1 := "PT801_VAL", in2 := "PT801_LOW")
      wire#w12
      Coil( "ALARM_PT801" )
   END_RUNG
   RUNG wire#powerrail
      Contact( "ALARM_PT801" )
      I_Contact( #CLEAR )
   END_RUNG wire#w12
   RUNG wire#powerrail
      { S7_Templates := "SrcType := Real" } GT_Contact(in1 := "PT901_VAL", in2 := "PT901_HIGH")
      wire#w13
      Coil( "ALARM_PT901" )
   END_RUNG
   RUNG wire#powerrail
      Contact( "ALARM_PT901" )
      I_Contact( #CLEAR )
   END_RUNG wire#w13
   RUNG wire#powerrail
      I_Contact( "ABORT_ON" )
      I_Contact( "STEP_0_ON" )
      I_Contact( "DOORS_CLOSED" )
      Contact( "AlwaysFALSE" )
      Coil( "ALARM_DOORS_OPEN" )
   END_RUNG
   // the same network as SCL:
   "ALARM_PT101" := ("PT101_VAL" < "PT101_LOW") OR ("ALARM_PT101" AND NOT #CLEAR);
   "ALARM_PT102" := ("PT102_VAL" > "PT102_HIGH") OR ("ALARM_PT102" AND NOT #CLEAR);
   "ALARM_PT201" := ("PT201_VAL" < "PT201_LOW_C") OR ("ALARM_PT201" AND NOT #CLEAR);
   "ALARM_PT202" := ("PT202_VAL" > "PT202_HIGH") OR ("ALARM_PT202" AND NOT #CLEAR);
   "ALARM_PT301" := ("PT301_VAL" < "PT301_LOW") OR ("ALARM_PT301" AND NOT #CLEAR);
   "ALARM_PT302" := ("PT302_VAL" > "PT302_HIGH") OR ("ALARM_PT302" AND NOT #CLEAR);
   "ALARM_PT401" := ("PT401_VAL" < "PT401_LOW") OR ("ALARM_PT401" AND NOT #CLEAR);